VERSION : 0.1
   VAR
      Line_A1_Save_Data : Bool;
      Line_A1_Save_Data_Advance : Bool;
      Line_A1_Start : Bool;
      Line_A1_Enable : Bool := 0;
      Line_A1_Conveyer_on_Time : Time := T#26MS;
      Line_A1_Conveyer_off_Time : Time := T#27MS;
      Line_A1_Sampling_Time : Time := T#28MS;
      Line_A1_Sampling_OpenTime : Time := T#29MS;
      Line_A1_Feeder_Intensity : Int := 30;
      Line_A1_Feeder_DelayTime : Time;
      Line_A1_Enable_Manual : Bool;
      Line_A1_Conveyor_Start_Manual : Bool;
      Line_A1_Big_Silo_Start_Manual : Bool;
      Line_A1_Below_Conveyor_Start_Manual : Bool;
      Line_A1_Feeder_Start_Manual : Bool;
      Line_A1_Sample_Start_Manual : Bool;
      Line_A1_Feeder_Delay_Before_Stop_Time : Time;
      Line_A1_Empty_Line_Time : Time;
      Line_A1_Big_Silo_Delay_Start : Time;
      Line_A1_Empty_Line : Bool;
      Line_A1_Feeder_Delay_After_Start_Time : Time;
      Line_A2_Save_Data : Bool;
      Line_A2_Save_Data_Advance : Bool;
      Line_A2_Start : Bool;
      Line_A2_Enable : Bool;
      Line_A2_Conveyer_on_Time : Time := T#8S_400MS;
      Line_A2_Conveyer_off_Time : Time := T#30s;
      Line_A2_Sampling_Time : Time := T#2M;
      Line_A2_Sampling_OpenTime : Time := T#9S_500MS;
      Line_A2_Feeder_Intensity : Int;
      Line_A2_Feeder_DelayTime : Time;
      Line_A2_Enable_Manual : Bool;
      Line_A2_Conveyor_Start_Manual : Bool;
      Line_A2_Big_Silo_Start_Manual : Bool;
      Line_A2_Below_Conveyor_Start_Manual : Bool;
      Line_A2_Feeder_Start_Manual : Bool;
      Line_A2_Sample_Start_Manual : Bool;
      Line_A2_Feeder_Delay_Before_Stop_Time : Time;
      Line_A2_Empty_Line_Time : Time;
      Line_A2_Big_Silo_Delay_Start : Time;
      Line_A2_Empty_Line : Bool;
      Line_A2_Feeder_Delay_After_Start_Time : Time;
      Line_B1_Save_Data : Bool;
      Line_B1_Save_Data_Advance : Bool;
      Line_B1_Start : Bool;
      Line_B1_Enable : Bool := 0;
      Line_B1_Conveyer_on_Time : Time := T#8S_400MS;
      Line_B1_Conveyer_off_Time : Time := T#30s;
      Line_B1_Sampling_Time : Time := T#2M;
      Line_B1_Sampling_OpenTime : Time := T#9S_500MS;
      Line_B1_Feeder_Intensity : Int;
      Line_B1_Feeder_DelayTime : Time;
      Line_B1_Enable_Manual : Bool;
      Line_B1_Conveyor_Start_Manual : Bool;
      Line_B1_Big_Silo_Start_Manual : Bool;
      Line_B1_Below_Conveyor_Start_Manual : Bool;
      Line_B1_Feeder_Start_Manual : Bool;
      Line_B1_Sample_Start_Manual : Bool;
      Line_B1_Feeder_Delay_Before_Stop_Time : Time;
      Line_B1_Empty_Line_Time : Time;
      Line_B1_Big_Silo_Delay_Start : Time;
      Line_B1_Empty_Line : Bool;
      Line_B1_Feeder_Delay_After_Start_Time : Time;
      Line_B2_Save_Data : Bool;
      Line_B2_Save_Data_Advance : Bool;
      Line_B2_Start : Bool;
      Line_B2_Enable : Bool := 0;
      Line_B2_Conveyer_on_Time : Time := T#8S_400MS;
      Line_B2_Conveyer_off_Time : Time := T#30s;
      Line_B2_Sampling_Time : Time := T#2M;
      Line_B2_Sampling_OpenTime : Time := T#9S_500MS;
      Line_B2_Feeder_Intensity : Int;
      Line_B2_Feeder_DelayTime : Time;
      Line_B2_Enable_Manual : Bool;
      Line_B2_Conveyor_Start_Manual : Bool;
      Line_B2_Big_Silo_Start_Manual : Bool;
      Line_B2_Below_Conveyor_Start_Manual : Bool;
      Line_B2_Feeder_Start_Manual : Bool;
      Line_B2_Sample_Start_Manual : Bool;
      Line_B2_Feeder_Delay_Before_Stop_Time : Time;
      Line_B2_Empty_Line_Time : Time;
      Line_B2_Big_Silo_Delay_Start : Time;
      Line_B2_Empty_Line : Bool;
      Line_B2_Feeder_Delay_After_Start_Time : Time;
      Conveyer_B3_Left : Bool;
   END_VAR
BEGIN
END_DATA_BLOCK

DATA_BLOCK "Empty Line A1 A2_DB"   // DB47
{ S7_Optimized_Access := 'TRUE' }
VERSION : 0.1
// stored: InstanceOfName Empty Line A1 A2
"Empty Line A1 A2"
BEGIN
END_DATA_BLOCK

DATA_BLOCK "Empty Line B1 B2_DB"   // DB48
{ S7_Optimized_Access := 'TRUE' }
VERSION : 0.1
// stored: InstanceOfName Empty Line B1 B2
"Empty Line B1 B2"
BEGIN
END_DATA_BLOCK

DATA_BLOCK "WebDataPrepaare_DB"   // DB49
{ S7_Optimized_Access := 'TRUE' }
VERSION : 0.1
// stored: InstanceOfName WebDataPrepaare
"WebDataPrepaare"
BEGIN
END_DATA_BLOCK

DATA_BLOCK "SaveDataToDataBlock A1_DB"   // DB51
{ S7_Optimized_Access := 'TRUE' }
VERSION : 0.1
// stored: InstanceOfName SaveDataToDataBlock A1
"SaveDataToDataBlock A1"
BEGIN
END_DATA_BLOCK

DATA_BLOCK "SaveDataToDataBlock A2_DB"   // DB52
{ S7_Optimized_Access := 'TRUE' }
VERSION : 0.1
// stored: InstanceOfName SaveDataToDataBlock A2
"SaveDataToDataBlock A2"
BEGIN
END_DATA_BLOCK

DATA_BLOCK "SaveDataToDataBlock B1_DB"   // DB53
{ S7_Optimized_Access := 'TRUE' }
VERSION : 0.1
// stored: InstanceOfName SaveDataToDataBlock B1
"SaveDataToDataBlock B1"
BEGIN
END_DATA_BLOCK

DATA_BLOCK "SaveDataToDataBlock B2_DB"   // DB54
{ S7_Optimized_Access := 'TRUE' }
VERSION : 0.1
// stored: InstanceOfName SaveDataToDataBlock B2
"SaveDataToDataBlock B2"
BEGIN
END_DATA_BLOCK

// folder: System blocks/Program resources

DATA_BLOCK "Timer_On_A1_Conveyer"   // DB6
{ S7_Optimized_Access := 'TRUE' }
AUTHOR : Simatic
FAMILY : IEC
NAME : IEC_TMR
VERSION : 1.0
// stored: InstanceOfName IEC_TIMER
"IEC_TIMER"
BEGIN
END_DATA_BLOCK

DATA_BLOCK "Timer_Off_A1_Conveyer"   // DB8
{ S7_Optimized_Access := 'TRUE' }
AUTHOR : Simatic
FAMILY : IEC
NAME : IEC_TMR
VERSION : 1.0
// stored: InstanceOfName IEC_TIMER
"IEC_TIMER"
BEGIN
END_DATA_BLOCK

DATA_BLOCK "Timer_On_A2_Conveyer"   // DB10
{ S7_Optimized_Access := 'TRUE' }
AUTHOR : Simatic
FAMILY : IEC
NAME : IEC_TMR
VERSION : 1.0
// stored: InstanceOfName IEC_TIMER
"IEC_TIMER"
BEGIN
END_DATA_BLOCK

DATA_BLOCK "Timer_Off_A2_Conveyer"   // DB11
{ S7_Optimized_Access := 'TRUE' }
AUTHOR : Simatic
FAMILY : IEC
NAME : IEC_TMR
VERSION : 1.0
// stored: InstanceOfName IEC_TIMER
"IEC_TIMER"
BEGIN
END_DATA_BLOCK

DATA_BLOCK "Timer_On_B1_Conveyer"   // DB14
{ S7_Optimized_Access := 'TRUE' }
AUTHOR : Simatic
FAMILY : IEC
NAME : IEC_TMR
VERSION : 1.0
// stored: InstanceOfName IEC_TIMER
"IEC_TIMER"
BEGIN
END_DATA_BLOCK

DATA_BLOCK "Timer_Off_B1_Conveyer"   // DB15
{ S7_Optimized_Access := 'TRUE' }
AUTHOR : Simatic
FAMILY : IEC
NAME : IEC_TMR
VERSION : 1.0
// stored: InstanceOfName IEC_TIMER
"IEC_TIMER"
BEGIN
END_DATA_BLOCK

DATA_BLOCK "Timer_On_B2_Conveyer"   // DB16
{ S7_Optimized_Access := 'TRUE' }
AUTHOR : Simatic
FAMILY : IEC
NAME : IEC_TMR
VERSION : 1.0
// stored: InstanceOfName IEC_TIMER
"IEC_TIMER"
BEGIN
END_DATA_BLOCK

DATA_BLOCK "Timer_Off_B2_Conveyer"   // DB24
{ S7_Optimized_Access := 'TRUE' }
AUTHOR : Simatic
FAMILY : IEC
NAME : IEC_TMR
VERSION : 1.0
// stored: InstanceOfName IEC_TIMER
"IEC_TIMER"
BEGIN
END_DATA_BLOCK

DATA_BLOCK "Timer_Before_On_Sample_A1"   // DB25
{ S7_Optimized_Access := 'TRUE' }
AUTHOR : Simatic
FAMILY : IEC
NAME : IEC_TMR
VERSION : 1.0
// stored: InstanceOfName IEC_TIMER
"IEC_TIMER"
BEGIN
END_DATA_BLOCK

DATA_BLOCK "Timer_Sample_Open_Time_A1"   // DB26
{ S7_Optimized_Access := 'TRUE' }
AUTHOR : Simatic
FAMILY : IEC
NAME : IEC_TMR
VERSION : 1.0
// stored: InstanceOfName IEC_TIMER
"IEC_TIMER"
BEGIN
END_DATA_BLOCK

DATA_BLOCK "Timer_Before_On_Sample_B1"   // DB27
{ S7_Optimized_Access := 'TRUE' }
AUTHOR : Simatic
FAMILY : IEC
NAME : IEC_TMR
VERSION : 1.0
// stored: InstanceOfName IEC_TIMER
"IEC_TIMER"
BEGIN
END_DATA_BLOCK

DATA_BLOCK "Timer_Before_On_Sample_A2"   // DB28
{ S7_Optimized_Access := 'TRUE' }
AUTHOR : Simatic
FAMILY : IEC
NAME : IEC_TMR
VERSION : 1.0
// stored: InstanceOfName IEC_TIMER
"IEC_TIMER"
BEGIN
END_DATA_BLOCK

DATA_BLOCK "Timer_Sample_Open_Time_B1"   // DB29
{ S7_Optimized_Access := 'TRUE' }
AUTHOR : Simatic
FAMILY : IEC
NAME : IEC_TMR
VERSION : 1.0
// stored: InstanceOfName IEC_TIMER
"IEC_TIMER"
BEGIN
END_DATA_BLOCK

DATA_BLOCK "Timer_Before_On_Sample_B2"   // DB30
{ S7_Optimized_Access := 'TRUE' }
AUTHOR : Simatic
FAMILY : IEC
NAME : IEC_TMR
VERSION : 1.0
// stored: InstanceOfName IEC_TIMER
"IEC_TIMER"
BEGIN
END_DATA_BLOCK

DATA_BLOCK "Timer_Sample_Open_Time_B2"   // DB31
{ S7_Optimized_Access := 'TRUE' }
AUTHOR : Simatic
FAMILY : IEC
NAME : IEC_TMR
VERSION : 1.0
// stored: InstanceOfName IEC_TIMER
"IEC_TIMER"
BEGIN
END_DATA_BLOCK

DATA_BLOCK "Timer_Sample_Open_Time_A2"   // DB35
{ S7_Optimized_Access := 'TRUE' }
AUTHOR : Simatic
FAMILY : IEC
NAME : IEC_TMR
VERSION : 1.0
// stored: InstanceOfName IEC_TIMER
"IEC_TIMER"
BEGIN
END_DATA_BLOCK

DATA_BLOCK "Timer_Silo_Big_B_Off_Time"   // DB36
{ S7_Optimized_Access := 'TRUE' }
AUTHOR : Simatic
FAMILY : IEC
NAME : IEC_TMR
VERSION : 1.0
// stored: InstanceOfName IEC_TIMER
"IEC_TIMER"
BEGIN
END_DATA_BLOCK

DATA_BLOCK "Timer_Silo_Big_A_Off_Time"   // DB37
{ S7_Optimized_Access := 'TRUE' }
AUTHOR : Simatic
FAMILY : IEC
NAME : IEC_TMR
VERSION : 1.0
// stored: InstanceOfName IEC_TIMER
"IEC_TIMER"
BEGIN
END_DATA_BLOCK

DATA_BLOCK "A1_Feeder_On_Delay_Timer"   // DB38
{ S7_Optimized_Access := 'TRUE' }
AUTHOR : Simatic
FAMILY : IEC
NAME : IEC_TMR
VERSION : 1.0
// stored: InstanceOfName IEC_TIMER
"IEC_TIMER"
BEGIN
END_DATA_BLOCK

DATA_BLOCK "A2_Feeder_On_Delay_Timer"   // DB39
{ S7_Optimized_Access := 'TRUE' }
AUTHOR : Simatic
FAMILY : IEC
NAME : IEC_TMR
VERSION : 1.0
// stored: InstanceOfName IEC_TIMER
"IEC_TIMER"
BEGIN
END_DATA_BLOCK

DATA_BLOCK "B1_Feeder_On_Delay_Timer"   // DB40
{ S7_Optimized_Access := 'TRUE' }
AUTHOR : Simatic
FAMILY : IEC
NAME : IEC_TMR
VERSION : 1.0
// stored: InstanceOfName IEC_TIMER
"IEC_TIMER"
BEGIN
END_DATA_BLOCK

DATA_BLOCK "B2_Feeder_On_Delay_Timer"   // DB41
{ S7_Optimized_Access := 'TRUE' }
AUTHOR : Simatic
FAMILY : IEC
NAME : IEC_TMR
VERSION : 1.0
// stored: InstanceOfName IEC_TIMER
"IEC_TIMER"
BEGIN
END_DATA_BLOCK

DATA_BLOCK "Timer_A1_Empty_Line_DB"   // DB42
{ S7_Optimized_Access := 'TRUE' }
AUTHOR : Simatic
FAMILY : IEC
NAME : IEC_TMR
VERSION : 1.0
// stored: InstanceOfName IEC_TIMER
"IEC_TIMER"
BEGIN
END_DATA_BLOCK

DATA_BLOCK "Timer_A2_Empty_Line_DB"   // DB43
{ S7_Optimized_Access := 'TRUE' }
AUTHOR : Simatic
FAMILY : IEC
NAME : IEC_TMR
VERSION : 1.0
// stored: InstanceOfName IEC_TIMER
"IEC_TIMER"
BEGIN
END_DATA_BLOCK

DATA_BLOCK "Timer_B1_Empty_Line_DB"   // DB44
{ S7_Optimized_Access := 'TRUE' }
AUTHOR : Simatic
FAMILY : IEC
NAME : IEC_TMR
VERSION : 1.0
// stored: InstanceOfName IEC_TIMER
"IEC_TIMER"
BEGIN
END_DATA_BLOCK

DATA_BLOCK "Timer_B2_Empty_Line_DB"   // DB46
{ S7_Optimized_Access := 'TRUE' }
AUTHOR : Simatic
FAMILY : IEC
NAME : IEC_TMR
VERSION : 1.0
// stored: InstanceOfName IEC_TIMER
"IEC_TIMER"
BEGIN
END_DATA_BLOCK

DATA_BLOCK "Timer_A1_Reset_Save_Data"   // DB50
{ S7_Optimized_Access := 'TRUE' }
AUTHOR : Simatic
FAMILY : IEC
NAME : IEC_TMR
VERSION : 1.0
// stored: InstanceOfName IEC_TIMER
"IEC_TIMER"
BEGIN
END_DATA_BLOCK

// folder: (top level)

FUNCTION_BLOCK "Conveyer A1"   // FB1, LAD
{ S7_Optimized_Access := 'TRUE' }
VERSION : 0.1
   VAR_TEMP   // added for the SCL form of the ladder/FBD networks
      _w1 : Bool;
   END_VAR
BEGIN

REGION Network 1: Run Consent Line A1
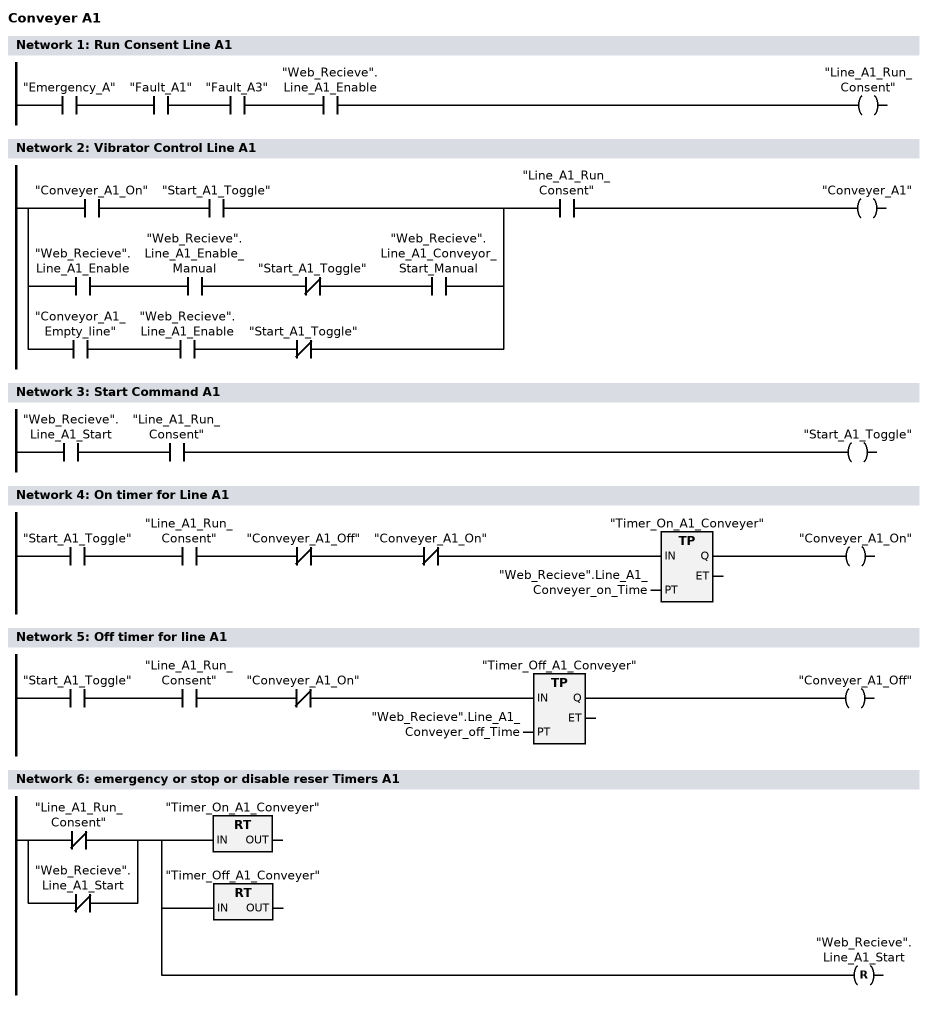
   RUNG wire#powerrail
      Contact( "Emergency_A" )
      Contact( "Fault_A1" )
      Contact( "Fault_A3" )
      Contact( "Web_Recieve".Line_A1_Enable )
      Coil( "Line_A1_Run_Consent" )
   END_RUNG
   // the same network as SCL:
   "Line_A1_Run_Consent" := "Emergency_A" AND "Fault_A1" AND "Fault_A3" AND "Web_Recieve".Line_A1_Enable;
END_REGION

REGION Network 2: Vibrator Control Line A1
   RUNG wire#powerrail
      Contact( "Conveyer_A1_On" )
      Contact( "Start_A1_Toggle" )
      wire#w1
      Contact( "Line_A1_Run_Consent" )
      Coil( "Conveyer_A1" )
   END_RUNG
   RUNG wire#powerrail
      Contact( "Web_Recieve".Line_A1_Enable )
      Contact( "Web_Recieve".Line_A1_Enable_Manual )
      I_Contact( "Start_A1_Toggle" )
      Contact( "Web_Recieve".Line_A1_Conveyor_Start_Manual )
   END_RUNG wire#w1
   RUNG wire#powerrail
      Contact( "Conveyor_A1_Empty_line" )
      Contact( "Web_Recieve".Line_A1_Enable )
      I_Contact( "Start_A1_Toggle" )
   END_RUNG wire#w1
   // the same network as SCL:
   "Conveyer_A1" := (("Conveyer_A1_On" AND "Start_A1_Toggle") OR ("Web_Recieve".Line_A1_Enable AND "Web_Recieve".Line_A1_Enable_Manual AND NOT "Start_A1_Toggle" AND "Web_Recieve".Line_A1_Conveyor_Start_Manual) OR ("Conveyor_A1_Empty_line" AND "Web_Recieve".Line_A1_Enable AND NOT "Start_A1_Toggle")) AND "Line_A1_Run_Consent";
END_REGION

REGION Network 3: Start Command A1
   RUNG wire#powerrail
      Contact( "Web_Recieve".Line_A1_Start )
      Contact( "Line_A1_Run_Consent" )
      Coil( "Start_A1_Toggle" )
   END_RUNG
   // the same network as SCL:
   "Start_A1_Toggle" := "Web_Recieve".Line_A1_Start AND "Line_A1_Run_Consent";
END_REGION

REGION Network 4: On timer for Line A1
   "Timer_On_A1_Conveyer".TP(IN := "Start_A1_Toggle" AND "Line_A1_Run_Consent" AND NOT "Conveyer_A1_Off" AND NOT "Conveyer_A1_On",
                           PT := "Web_Recieve".Line_A1_Conveyer_on_Time);
   "Conveyer_A1_On" := "Timer_On_A1_Conveyer".Q;
END_REGION

REGION Network 5: Off timer for line A1
   "Timer_Off_A1_Conveyer".TP(IN := "Start_A1_Toggle" AND "Line_A1_Run_Consent" AND NOT "Conveyer_A1_On",
                           PT := "Web_Recieve".Line_A1_Conveyer_off_Time);
   "Conveyer_A1_Off" := "Timer_Off_A1_Conveyer".Q;
END_REGION

REGION Network 6: emergency or stop or disable reser Timers A1
   RUNG wire#powerrail
      I_Contact( "Line_A1_Run_Consent" )
      wire#w1
      RT_Coil( "Timer_On_A1_Conveyer" )
   END_RUNG
   RUNG wire#powerrail
      I_Contact( "Web_Recieve".Line_A1_Start )
   END_RUNG wire#w1
   RUNG wire#w1
      RT_Coil( "Timer_Off_A1_Conveyer" )
   END_RUNG
   RUNG wire#w1
      R_Coil( "Web_Recieve".Line_A1_Start )
   END_RUNG
   // the same network as SCL:
   #_w1 := NOT "Line_A1_Run_Consent" OR NOT "Web_Recieve".Line_A1_Start;
   IF #_w1 THEN
       RESET_TIMER("Timer_On_A1_Conveyer");
       RESET_TIMER("Timer_Off_A1_Conveyer");
       "Web_Recieve".Line_A1_Start := FALSE;
   END_IF;
END_REGION
END_FUNCTION_BLOCK

FUNCTION_BLOCK "Conveyer A2"   // FB2, LAD
{ S7_Optimized_Access := 'TRUE' }
VERSION : 0.1
   VAR_TEMP   // added for the SCL form of the ladder/FBD networks
      _w1 : Bool;
   END_VAR
BEGIN

REGION Network 1: Run Consent Line A2
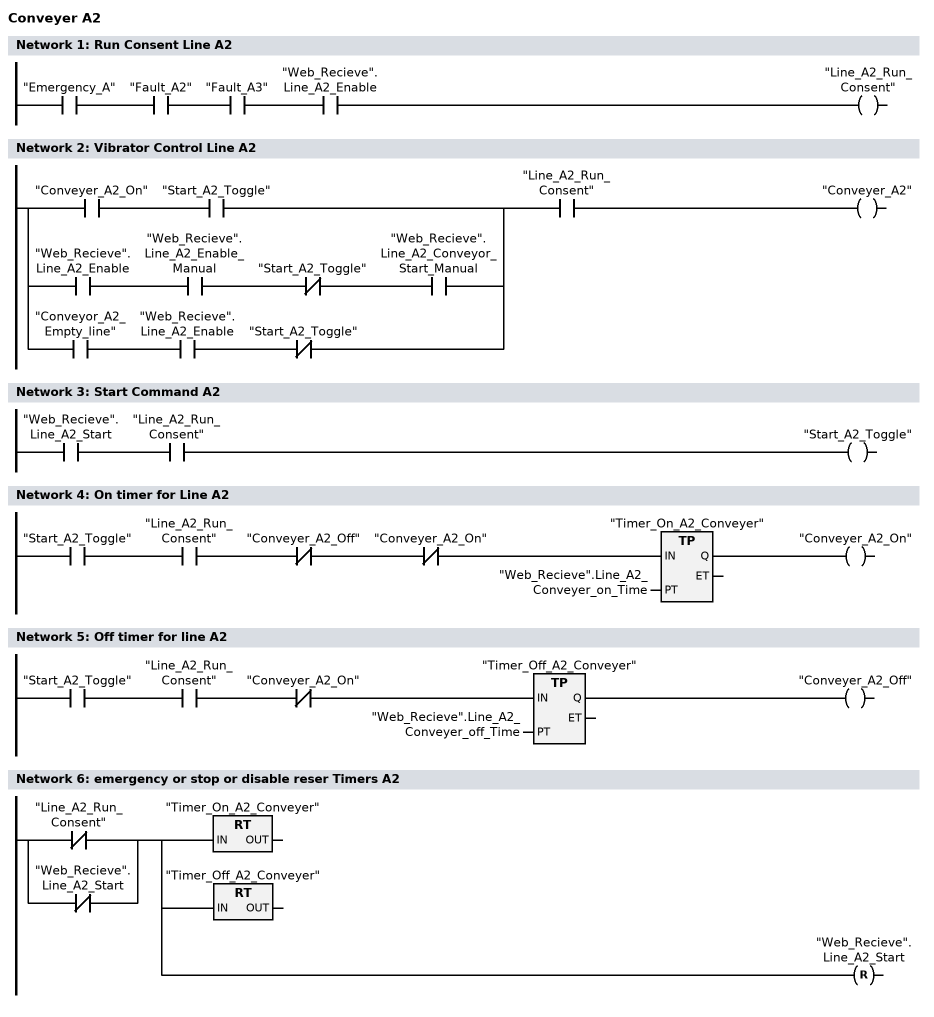
   RUNG wire#powerrail
      Contact( "Emergency_A" )
      Contact( "Fault_A2" )
      Contact( "Fault_A3" )
      Contact( "Web_Recieve".Line_A2_Enable )
      Coil( "Line_A2_Run_Consent" )
   END_RUNG
   // the same network as SCL:
   "Line_A2_Run_Consent" := "Emergency_A" AND "Fault_A2" AND "Fault_A3" AND "Web_Recieve".Line_A2_Enable;
END_REGION

REGION Network 2: Vibrator Control Line A2
   RUNG wire#powerrail
      Contact( "Conveyer_A2_On" )
      Contact( "Start_A2_Toggle" )
      wire#w1
      Contact( "Line_A2_Run_Consent" )
      Coil( "Conveyer_A2" )
   END_RUNG
   RUNG wire#powerrail
      Contact( "Web_Recieve".Line_A2_Enable )
      Contact( "Web_Recieve".Line_A2_Enable_Manual )
      I_Contact( "Start_A2_Toggle" )
      Contact( "Web_Recieve".Line_A2_Conveyor_Start_Manual )
   END_RUNG wire#w1
   RUNG wire#powerrail
      Contact( "Conveyor_A2_Empty_line" )
      Contact( "Web_Recieve".Line_A2_Enable )
      I_Contact( "Start_A2_Toggle" )
   END_RUNG wire#w1
   // the same network as SCL:
   "Conveyer_A2" := (("Conveyer_A2_On" AND "Start_A2_Toggle") OR ("Web_Recieve".Line_A2_Enable AND "Web_Recieve".Line_A2_Enable_Manual AND NOT "Start_A2_Toggle" AND "Web_Recieve".Line_A2_Conveyor_Start_Manual) OR ("Conveyor_A2_Empty_line" AND "Web_Recieve".Line_A2_Enable AND NOT "Start_A2_Toggle")) AND "Line_A2_Run_Consent";
END_REGION

REGION Network 3: Start Command A2
   RUNG wire#powerrail
      Contact( "Web_Recieve".Line_A2_Start )
      Contact( "Line_A2_Run_Consent" )
      Coil( "Start_A2_Toggle" )
   END_RUNG
   // the same network as SCL:
   "Start_A2_Toggle" := "Web_Recieve".Line_A2_Start AND "Line_A2_Run_Consent";
END_REGION

REGION Network 4: On timer for Line A2
   "Timer_On_A2_Conveyer".TP(IN := "Start_A2_Toggle" AND "Line_A2_Run_Consent" AND NOT "Conveyer_A2_Off" AND NOT "Conveyer_A2_On",
                           PT := "Web_Recieve".Line_A2_Conveyer_on_Time);
   "Conveyer_A2_On" := "Timer_On_A2_Conveyer".Q;
END_REGION

REGION Network 5: Off timer for line A2
   "Timer_Off_A2_Conveyer".TP(IN := "Start_A2_Toggle" AND "Line_A2_Run_Consent" AND NOT "Conveyer_A2_On",
                           PT := "Web_Recieve".Line_A2_Conveyer_off_Time);
   "Conveyer_A2_Off" := "Timer_Off_A2_Conveyer".Q;
END_REGION

REGION Network 6: emergency or stop or disable reser Timers A2
   RUNG wire#powerrail
      I_Contact( "Line_A2_Run_Consent" )
      wire#w1
      RT_Coil( "Timer_On_A2_Conveyer" )
   END_RUNG
   RUNG wire#powerrail
      I_Contact( "Web_Recieve".Line_A2_Start )
   END_RUNG wire#w1
   RUNG wire#w1
      RT_Coil( "Timer_Off_A2_Conveyer" )
   END_RUNG
   RUNG wire#w1
      R_Coil( "Web_Recieve".Line_A2_Start )
   END_RUNG
   // the same network as SCL:
   #_w1 := NOT "Line_A2_Run_Consent" OR NOT "Web_Recieve".Line_A2_Start;
   IF #_w1 THEN
       RESET_TIMER("Timer_On_A2_Conveyer");
       RESET_TIMER("Timer_Off_A2_Conveyer");
       "Web_Recieve".Line_A2_Start := FALSE;
   END_IF;
END_REGION
END_FUNCTION_BLOCK

FUNCTION_BLOCK "Conveyer B1"   // FB3, LAD
{ S7_Optimized_Access := 'TRUE' }
VERSION : 0.1
   VAR_TEMP   // added for the SCL form of the ladder/FBD networks
      _w1 : Bool;
      _w2 : Bool;
   END_VAR
BEGIN

REGION Network 1: Start Consent line A1
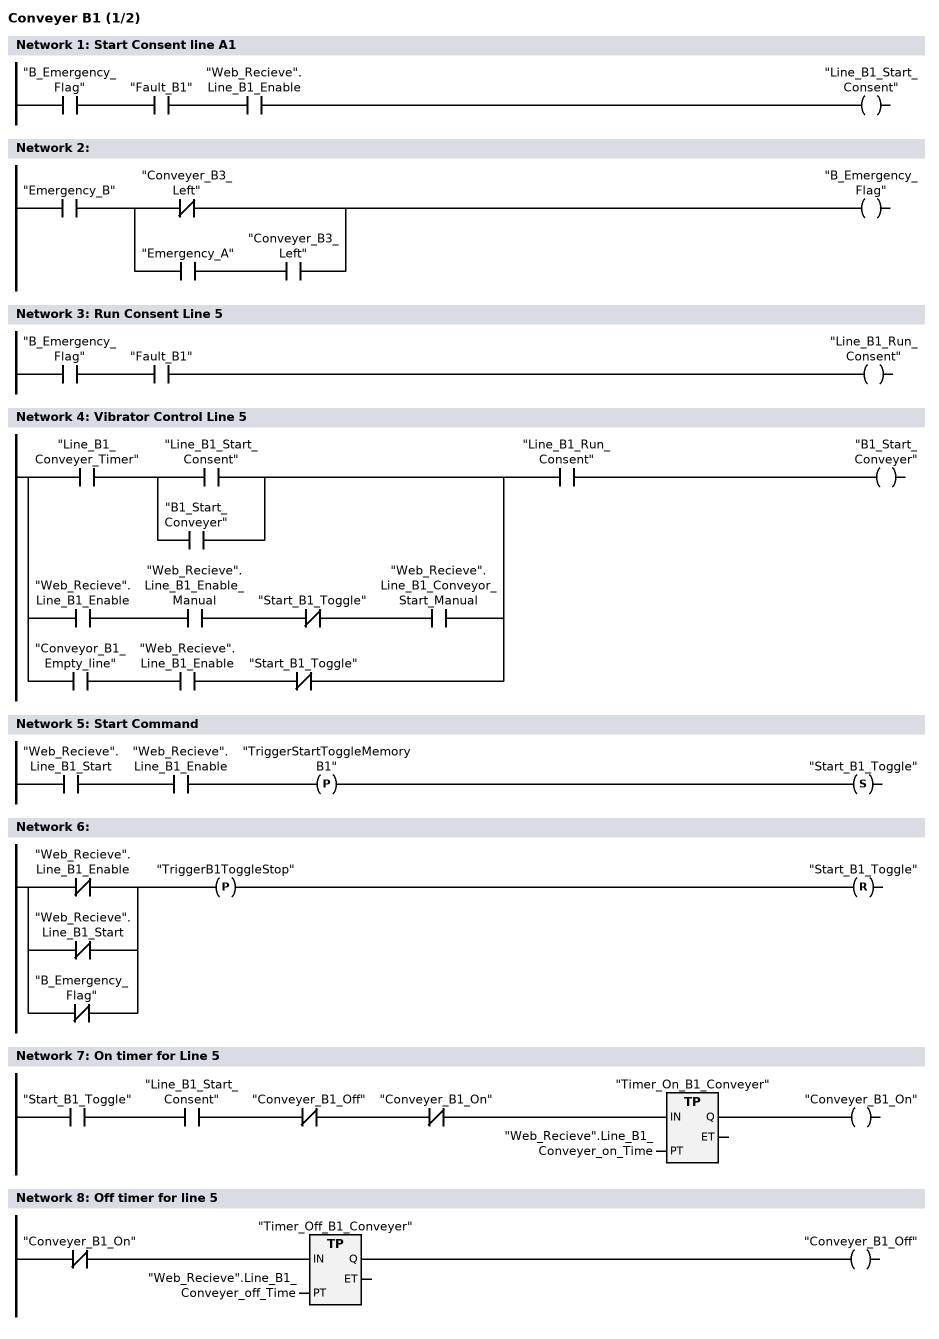
   RUNG wire#powerrail
      Contact( "B_Emergency_Flag" )
      Contact( "Fault_B1" )
      Contact( "Web_Recieve".Line_B1_Enable )
      Coil( "Line_B1_Start_Consent" )
   END_RUNG
   // the same network as SCL:
   "Line_B1_Start_Consent" := "B_Emergency_Flag" AND "Fault_B1" AND "Web_Recieve".Line_B1_Enable;
END_REGION

REGION Network 2
   RUNG wire#powerrail
      Contact( "Emergency_B" )
      wire#w1
      I_Contact( "Conveyer_B3_Left" )
      wire#w2
      Coil( "B_Emergency_Flag" )
   END_RUNG
   RUNG wire#w1
      Contact( "Emergency_A" )
      Contact( "Conveyer_B3_Left" )
   END_RUNG wire#w2
   // the same network as SCL:
   "B_Emergency_Flag" := "Emergency_B" AND (NOT "Conveyer_B3_Left" OR ("Emergency_A" AND "Conveyer_B3_Left"));
END_REGION

REGION Network 3: Run Consent Line 5
   RUNG wire#powerrail
      Contact( "B_Emergency_Flag" )
      Contact( "Fault_B1" )
      Coil( "Line_B1_Run_Consent" )
   END_RUNG
   // the same network as SCL:
   "Line_B1_Run_Consent" := "B_Emergency_Flag" AND "Fault_B1";
END_REGION

REGION Network 4: Vibrator Control Line 5
   RUNG wire#powerrail
      Contact( "Line_B1_Conveyer_Timer" )
      wire#w1
      Contact( "Line_B1_Start_Consent" )
      wire#w2
      Contact( "Line_B1_Run_Consent" )
      Coil( "B1_Start_Conveyer" )
   END_RUNG
   RUNG wire#w1
      Contact( "B1_Start_Conveyer" )
   END_RUNG wire#w2
   RUNG wire#powerrail
      Contact( "Web_Recieve".Line_B1_Enable )
      Contact( "Web_Recieve".Line_B1_Enable_Manual )
      I_Contact( "Start_B1_Toggle" )
      Contact( "Web_Recieve".Line_B1_Conveyor_Start_Manual )
   END_RUNG wire#w2
   RUNG wire#powerrail
      Contact( "Conveyor_B1_Empty_line" )
      Contact( "Web_Recieve".Line_B1_Enable )
      I_Contact( "Start_B1_Toggle" )
   END_RUNG wire#w2
   // the same network as SCL:
   "B1_Start_Conveyer" := (("Line_B1_Conveyer_Timer" AND ("Line_B1_Start_Consent" OR "B1_Start_Conveyer")) OR ("Web_Recieve".Line_B1_Enable AND "Web_Recieve".Line_B1_Enable_Manual AND NOT "Start_B1_Toggle" AND "Web_Recieve".Line_B1_Conveyor_Start_Manual) OR ("Conveyor_B1_Empty_line" AND "Web_Recieve".Line_B1_Enable AND NOT "Start_B1_Toggle")) AND "Line_B1_Run_Consent";
END_REGION

REGION Network 5: Start Command
   RUNG wire#powerrail
      Contact( "Web_Recieve".Line_B1_Start )
      Contact( "Web_Recieve".Line_B1_Enable )
      P_Trig( "TriggerStartToggleMemoryB1" )
      S_Coil( "Start_B1_Toggle" )
   END_RUNG
   // the same network as SCL:
   #_w1 := "Web_Recieve".Line_B1_Start AND "Web_Recieve".Line_B1_Enable;
   #_w2 := #_w1 AND NOT "TriggerStartToggleMemoryB1";   // rising edge
   "TriggerStartToggleMemoryB1" := #_w1;
   IF #_w2 THEN "Start_B1_Toggle" := TRUE; END_IF;
END_REGION

REGION Network 6
   RUNG wire#powerrail
      I_Contact( "Web_Recieve".Line_B1_Enable )
      wire#w1
      P_Trig( "TriggerB1ToggleStop" )
      R_Coil( "Start_B1_Toggle" )
   END_RUNG
   RUNG wire#powerrail
      I_Contact( "Web_Recieve".Line_B1_Start )
   END_RUNG wire#w1
   RUNG wire#powerrail
      I_Contact( "B_Emergency_Flag" )
   END_RUNG wire#w1
   // the same network as SCL:
   #_w1 := NOT "Web_Recieve".Line_B1_Enable OR NOT "Web_Recieve".Line_B1_Start OR NOT "B_Emergency_Flag";
   #_w2 := #_w1 AND NOT "TriggerB1ToggleStop";   // rising edge
   "TriggerB1ToggleStop" := #_w1;
   IF #_w2 THEN "Start_B1_Toggle" := FALSE; END_IF;
END_REGION

REGION Network 7: On timer for Line 5
   "Timer_On_B1_Conveyer".TP(IN := "Start_B1_Toggle" AND "Line_B1_Start_Consent" AND NOT "Conveyer_B1_Off" AND NOT "Conveyer_B1_On",
                           PT := "Web_Recieve".Line_B1_Conveyer_on_Time);
   "Conveyer_B1_On" := "Timer_On_B1_Conveyer".Q;
END_REGION

REGION Network 8: Off timer for line 5
   "Timer_Off_B1_Conveyer".TP(IN := NOT "Conveyer_B1_On", PT := "Web_Recieve".Line_B1_Conveyer_off_Time);
   "Conveyer_B1_Off" := "Timer_Off_B1_Conveyer".Q;
END_REGION

REGION Network 9
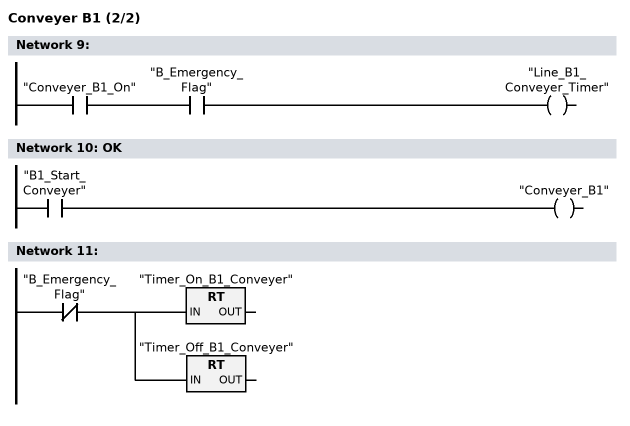
   RUNG wire#powerrail
      Contact( "Conveyer_B1_On" )
      Contact( "B_Emergency_Flag" )
      Coil( "Line_B1_Conveyer_Timer" )
   END_RUNG
   // the same network as SCL:
   "Line_B1_Conveyer_Timer" := "Conveyer_B1_On" AND "B_Emergency_Flag";
END_REGION

REGION Network 10: OK
   RUNG wire#powerrail
      Contact( "B1_Start_Conveyer" )
      Coil( "Conveyer_B1" )
   END_RUNG
   // the same network as SCL:
   "Conveyer_B1" := "B1_Start_Conveyer";
END_REGION

REGION Network 11
   RUNG wire#powerrail
      I_Contact( "B_Emergency_Flag" )
      wire#w1
      RT_Coil( "Timer_On_B1_Conveyer" )
   END_RUNG
   RUNG wire#w1
      RT_Coil( "Timer_Off_B1_Conveyer" )
   END_RUNG
   // the same network as SCL:
   IF NOT "B_Emergency_Flag" THEN
       RESET_TIMER("Timer_On_B1_Conveyer");
       RESET_TIMER("Timer_Off_B1_Conveyer");
   END_IF;
END_REGION
END_FUNCTION_BLOCK

FUNCTION_BLOCK "Conveyer B2"   // FB4, LAD
{ S7_Optimized_Access := 'TRUE' }
VERSION : 0.1
   VAR_TEMP   // added for the SCL form of the ladder/FBD networks
      _w1 : Bool;
      _w2 : Bool;
   END_VAR
BEGIN

REGION Network 1: Start Consent line A1
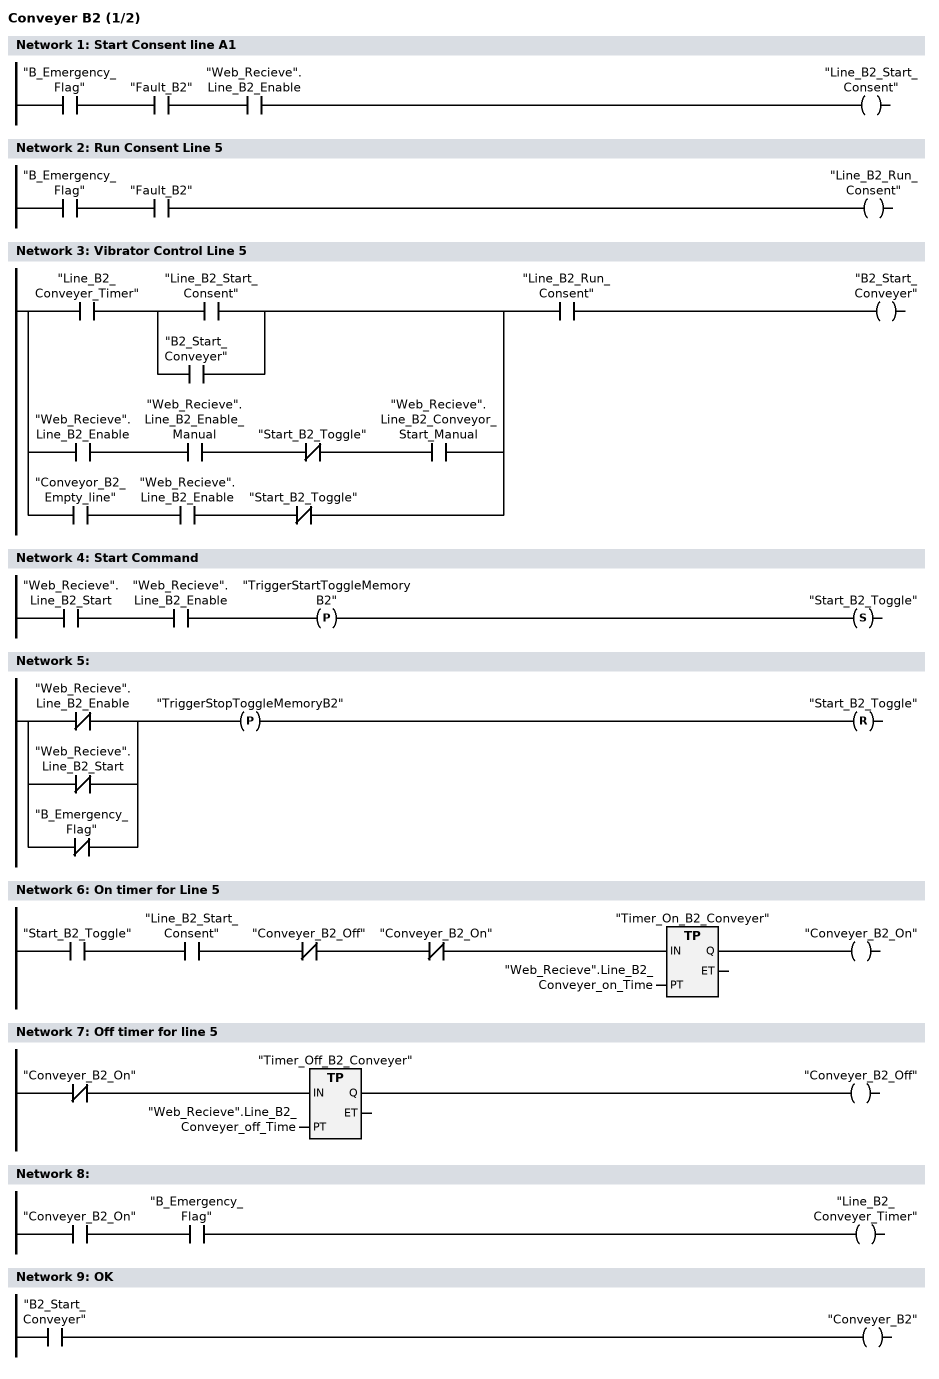
   RUNG wire#powerrail
      Contact( "B_Emergency_Flag" )
      Contact( "Fault_B2" )
      Contact( "Web_Recieve".Line_B2_Enable )
      Coil( "Line_B2_Start_Consent" )
   END_RUNG
   // the same network as SCL:
   "Line_B2_Start_Consent" := "B_Emergency_Flag" AND "Fault_B2" AND "Web_Recieve".Line_B2_Enable;
END_REGION

REGION Network 2: Run Consent Line 5
   RUNG wire#powerrail
      Contact( "B_Emergency_Flag" )
      Contact( "Fault_B2" )
      Coil( "Line_B2_Run_Consent" )
   END_RUNG
   // the same network as SCL:
   "Line_B2_Run_Consent" := "B_Emergency_Flag" AND "Fault_B2";
END_REGION

REGION Network 3: Vibrator Control Line 5
   RUNG wire#powerrail
      Contact( "Line_B2_Conveyer_Timer" )
      wire#w1
      Contact( "Line_B2_Start_Consent" )
      wire#w2
      Contact( "Line_B2_Run_Consent" )
      Coil( "B2_Start_Conveyer" )
   END_RUNG
   RUNG wire#w1
      Contact( "B2_Start_Conveyer" )
   END_RUNG wire#w2
   RUNG wire#powerrail
      Contact( "Web_Recieve".Line_B2_Enable )
      Contact( "Web_Recieve".Line_B2_Enable_Manual )
      I_Contact( "Start_B2_Toggle" )
      Contact( "Web_Recieve".Line_B2_Conveyor_Start_Manual )
   END_RUNG wire#w2
   RUNG wire#powerrail
      Contact( "Conveyor_B2_Empty_line" )
      Contact( "Web_Recieve".Line_B2_Enable )
      I_Contact( "Start_B2_Toggle" )
   END_RUNG wire#w2
   // the same network as SCL:
   "B2_Start_Conveyer" := (("Line_B2_Conveyer_Timer" AND ("Line_B2_Start_Consent" OR "B2_Start_Conveyer")) OR ("Web_Recieve".Line_B2_Enable AND "Web_Recieve".Line_B2_Enable_Manual AND NOT "Start_B2_Toggle" AND "Web_Recieve".Line_B2_Conveyor_Start_Manual) OR ("Conveyor_B2_Empty_line" AND "Web_Recieve".Line_B2_Enable AND NOT "Start_B2_Toggle")) AND "Line_B2_Run_Consent";
END_REGION

REGION Network 4: Start Command
   RUNG wire#powerrail
      Contact( "Web_Recieve".Line_B2_Start )
      Contact( "Web_Recieve".Line_B2_Enable )
      P_Trig( "TriggerStartToggleMemoryB2" )
      S_Coil( "Start_B2_Toggle" )
   END_RUNG
   // the same network as SCL:
   #_w1 := "Web_Recieve".Line_B2_Start AND "Web_Recieve".Line_B2_Enable;
   #_w2 := #_w1 AND NOT "TriggerStartToggleMemoryB2";   // rising edge
   "TriggerStartToggleMemoryB2" := #_w1;
   IF #_w2 THEN "Start_B2_Toggle" := TRUE; END_IF;
END_REGION

REGION Network 5
   RUNG wire#powerrail
      I_Contact( "Web_Recieve".Line_B2_Enable )
      wire#w1
      P_Trig( "TriggerStopToggleMemoryB2" )
      R_Coil( "Start_B2_Toggle" )
   END_RUNG
   RUNG wire#powerrail
      I_Contact( "Web_Recieve".Line_B2_Start )
   END_RUNG wire#w1
   RUNG wire#powerrail
      I_Contact( "B_Emergency_Flag" )
   END_RUNG wire#w1
   // the same network as SCL:
   #_w1 := NOT "Web_Recieve".Line_B2_Enable OR NOT "Web_Recieve".Line_B2_Start OR NOT "B_Emergency_Flag";
   #_w2 := #_w1 AND NOT "TriggerStopToggleMemoryB2";   // rising edge
   "TriggerStopToggleMemoryB2" := #_w1;
   IF #_w2 THEN "Start_B2_Toggle" := FALSE; END_IF;
END_REGION

REGION Network 6: On timer for Line 5
   "Timer_On_B2_Conveyer".TP(IN := "Start_B2_Toggle" AND "Line_B2_Start_Consent" AND NOT "Conveyer_B2_Off" AND NOT "Conveyer_B2_On",
                           PT := "Web_Recieve".Line_B2_Conveyer_on_Time);
   "Conveyer_B2_On" := "Timer_On_B2_Conveyer".Q;
END_REGION

REGION Network 7: Off timer for line 5
   "Timer_Off_B2_Conveyer".TP(IN := NOT "Conveyer_B2_On", PT := "Web_Recieve".Line_B2_Conveyer_off_Time);
   "Conveyer_B2_Off" := "Timer_Off_B2_Conveyer".Q;
END_REGION

REGION Network 8
   RUNG wire#powerrail
      Contact( "Conveyer_B2_On" )
      Contact( "B_Emergency_Flag" )
      Coil( "Line_B2_Conveyer_Timer" )
   END_RUNG
   // the same network as SCL:
   "Line_B2_Conveyer_Timer" := "Conveyer_B2_On" AND "B_Emergency_Flag";
END_REGION

REGION Network 9: OK
   RUNG wire#powerrail
      Contact( "B2_Start_Conveyer" )
      Coil( "Conveyer_B2" )
   END_RUNG
   // the same network as SCL:
   "Conveyer_B2" := "B2_Start_Conveyer";
END_REGION

REGION Network 10
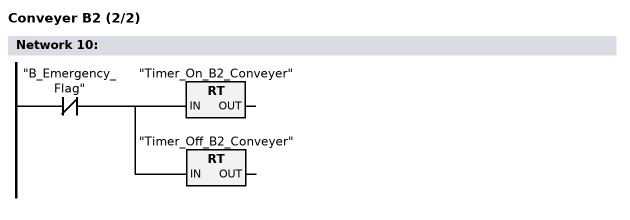
   RUNG wire#powerrail
      I_Contact( "B_Emergency_Flag" )
      wire#w1
      RT_Coil( "Timer_On_B2_Conveyer" )
   END_RUNG
   RUNG wire#w1
      RT_Coil( "Timer_Off_B2_Conveyer" )
   END_RUNG
   // the same network as SCL:
   IF NOT "B_Emergency_Flag" THEN
       RESET_TIMER("Timer_On_B2_Conveyer");
       RESET_TIMER("Timer_Off_B2_Conveyer");
   END_IF;
END_REGION
END_FUNCTION_BLOCK

FUNCTION_BLOCK "Vibrator A1"   // FB5, LAD
{ S7_Optimized_Access := 'TRUE' }
VERSION : 0.1
   VAR_TEMP
      RemainTime : DInt;
   END_VAR
BEGIN

REGION Network 1: Vibrator On Auto / Manual
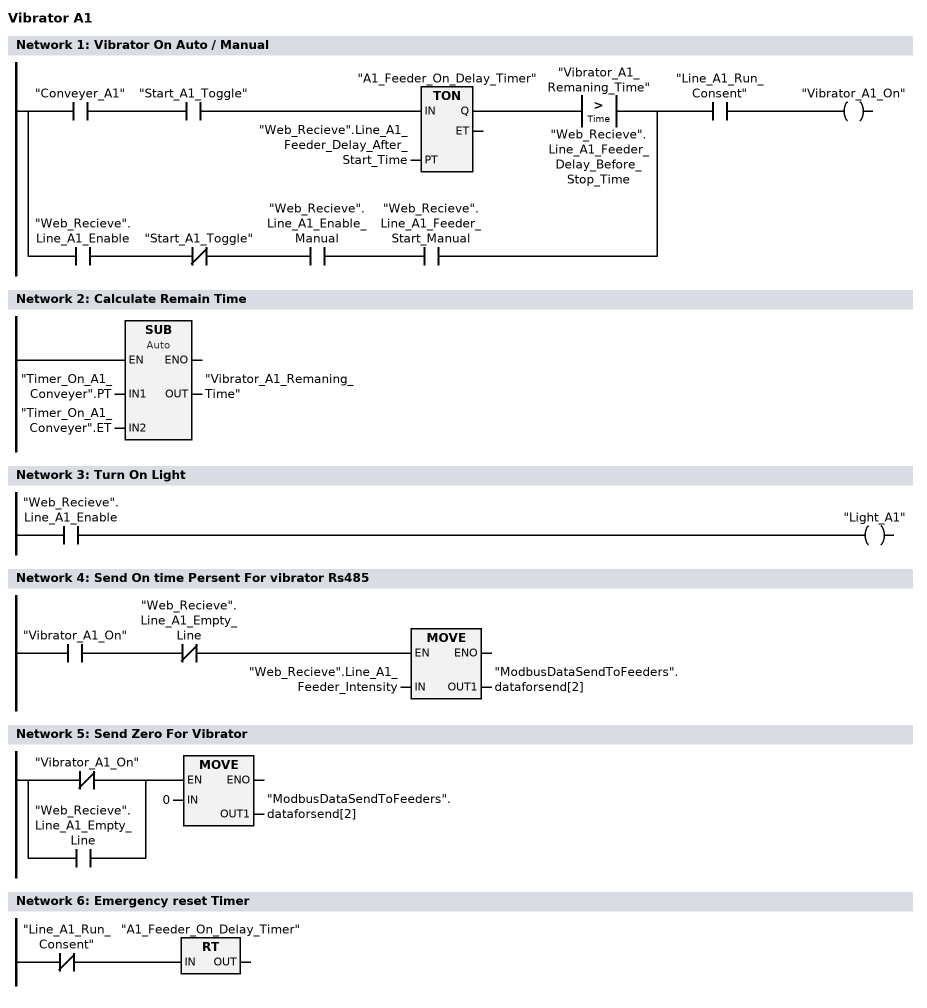
   "A1_Feeder_On_Delay_Timer".TON(IN := "Conveyer_A1" AND "Start_A1_Toggle",
                           PT := "Web_Recieve".Line_A1_Feeder_Delay_After_Start_Time);
   "Vibrator_A1_On" := (("A1_Feeder_On_Delay_Timer".Q AND ("Vibrator_A1_Remaning_Time" > "Web_Recieve".Line_A1_Feeder_Delay_Before_Stop_Time)) OR ("Web_Recieve".Line_A1_Enable AND NOT "Start_A1_Toggle" AND "Web_Recieve".Line_A1_Enable_Manual AND "Web_Recieve".Line_A1_Feeder_Start_Manual)) AND "Line_A1_Run_Consent";
END_REGION

REGION Network 2: Calculate Remain Time
   RUNG wire#powerrail
      Sub(in1 := "Timer_On_A1_Conveyer".PT, in2 := "Timer_On_A1_Conveyer".ET, out => "Vibrator_A1_Remaning_Time")
   END_RUNG
   // the same network as SCL:
   "Vibrator_A1_Remaning_Time" := "Timer_On_A1_Conveyer".PT - "Timer_On_A1_Conveyer".ET;
END_REGION

REGION Network 3: Turn On Light
   RUNG wire#powerrail
      Contact( "Web_Recieve".Line_A1_Enable )
      Coil( "Light_A1" )
   END_RUNG
   // the same network as SCL:
   "Light_A1" := "Web_Recieve".Line_A1_Enable;
END_REGION

REGION Network 4: Send On time Persent For vibrator Rs485
   RUNG wire#powerrail
      Contact( "Vibrator_A1_On" )
      I_Contact( "Web_Recieve".Line_A1_Empty_Line )
      Move(in := "Web_Recieve".Line_A1_Feeder_Intensity, out1 => "ModbusDataSendToFeeders".dataforsend[2])
   END_RUNG
   // the same network as SCL:
   IF "Vibrator_A1_On" AND NOT "Web_Recieve".Line_A1_Empty_Line THEN
       "ModbusDataSendToFeeders".dataforsend[2] := "Web_Recieve".Line_A1_Feeder_Intensity;
   END_IF;
END_REGION

REGION Network 5: Send Zero For Vibrator
   RUNG wire#powerrail
      I_Contact( "Vibrator_A1_On" )
      wire#w1
      Move(in := 0, out1 => "ModbusDataSendToFeeders".dataforsend[2])
   END_RUNG
   RUNG wire#powerrail
      Contact( "Web_Recieve".Line_A1_Empty_Line )
   END_RUNG wire#w1
   // the same network as SCL:
   IF NOT "Vibrator_A1_On" OR "Web_Recieve".Line_A1_Empty_Line THEN
       "ModbusDataSendToFeeders".dataforsend[2] := 0;
   END_IF;
END_REGION

REGION Network 6: Emergency reset Timer
   RUNG wire#powerrail
      I_Contact( "Line_A1_Run_Consent" )
      RT_Coil( "A1_Feeder_On_Delay_Timer" )
   END_RUNG
   // the same network as SCL:
   IF NOT "Line_A1_Run_Consent" THEN RESET_TIMER("A1_Feeder_On_Delay_Timer"); END_IF;
END_REGION
END_FUNCTION_BLOCK

FUNCTION_BLOCK "Vibrator A2"   // FB6, LAD
{ S7_Optimized_Access := 'TRUE' }
VERSION : 0.1
   VAR_TEMP
      RemainTime : DInt;
   END_VAR
BEGIN

REGION Network 1: Vibrator On Auto / Manual
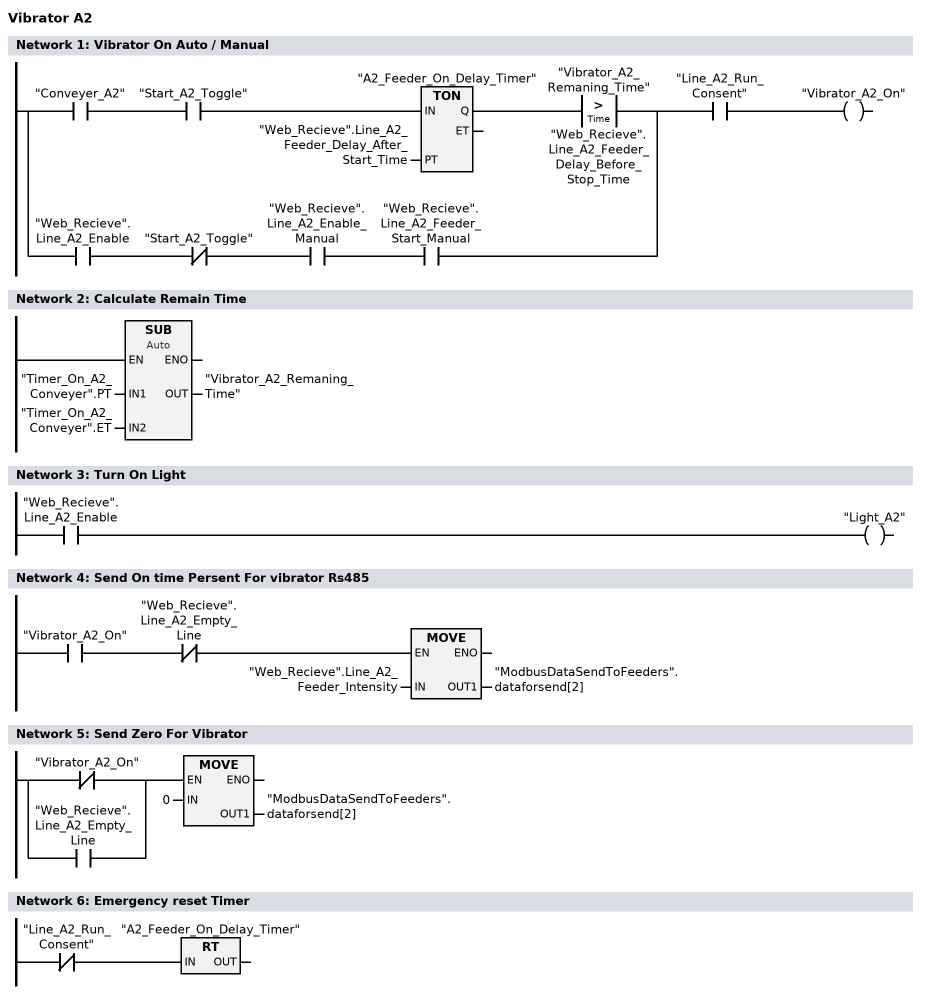
   "A2_Feeder_On_Delay_Timer".TON(IN := "Conveyer_A2" AND "Start_A2_Toggle",
                           PT := "Web_Recieve".Line_A2_Feeder_Delay_After_Start_Time);
   "Vibrator_A2_On" := (("A2_Feeder_On_Delay_Timer".Q AND ("Vibrator_A2_Remaning_Time" > "Web_Recieve".Line_A2_Feeder_Delay_Before_Stop_Time)) OR ("Web_Recieve".Line_A2_Enable AND NOT "Start_A2_Toggle" AND "Web_Recieve".Line_A2_Enable_Manual AND "Web_Recieve".Line_A2_Feeder_Start_Manual)) AND "Line_A2_Run_Consent";
END_REGION

REGION Network 2: Calculate Remain Time
   RUNG wire#powerrail
      Sub(in1 := "Timer_On_A2_Conveyer".PT, in2 := "Timer_On_A2_Conveyer".ET, out => "Vibrator_A2_Remaning_Time")
   END_RUNG
   // the same network as SCL:
   "Vibrator_A2_Remaning_Time" := "Timer_On_A2_Conveyer".PT - "Timer_On_A2_Conveyer".ET;
END_REGION

REGION Network 3: Turn On Light
   RUNG wire#powerrail
      Contact( "Web_Recieve".Line_A2_Enable )
      Coil( "Light_A2" )
   END_RUNG
   // the same network as SCL:
   "Light_A2" := "Web_Recieve".Line_A2_Enable;
END_REGION

REGION Network 4: Send On time Persent For vibrator Rs485
   RUNG wire#powerrail
      Contact( "Vibrator_A2_On" )
      I_Contact( "Web_Recieve".Line_A2_Empty_Line )
      Move(in := "Web_Recieve".Line_A2_Feeder_Intensity, out1 => "ModbusDataSendToFeeders".dataforsend[2])
   END_RUNG
   // the same network as SCL:
   IF "Vibrator_A2_On" AND NOT "Web_Recieve".Line_A2_Empty_Line THEN
       "ModbusDataSendToFeeders".dataforsend[2] := "Web_Recieve".Line_A2_Feeder_Intensity;
   END_IF;
END_REGION

REGION Network 5: Send Zero For Vibrator
   RUNG wire#powerrail
      I_Contact( "Vibrator_A2_On" )
      wire#w1
      Move(in := 0, out1 => "ModbusDataSendToFeeders".dataforsend[2])
   END_RUNG
   RUNG wire#powerrail
      Contact( "Web_Recieve".Line_A2_Empty_Line )
   END_RUNG wire#w1
   // the same network as SCL:
   IF NOT "Vibrator_A2_On" OR "Web_Recieve".Line_A2_Empty_Line THEN
       "ModbusDataSendToFeeders".dataforsend[2] := 0;
   END_IF;
END_REGION

REGION Network 6: Emergency reset Timer
   RUNG wire#powerrail
      I_Contact( "Line_A2_Run_Consent" )
      RT_Coil( "A2_Feeder_On_Delay_Timer" )
   END_RUNG
   // the same network as SCL:
   IF NOT "Line_A2_Run_Consent" THEN RESET_TIMER("A2_Feeder_On_Delay_Timer"); END_IF;
END_REGION
END_FUNCTION_BLOCK

